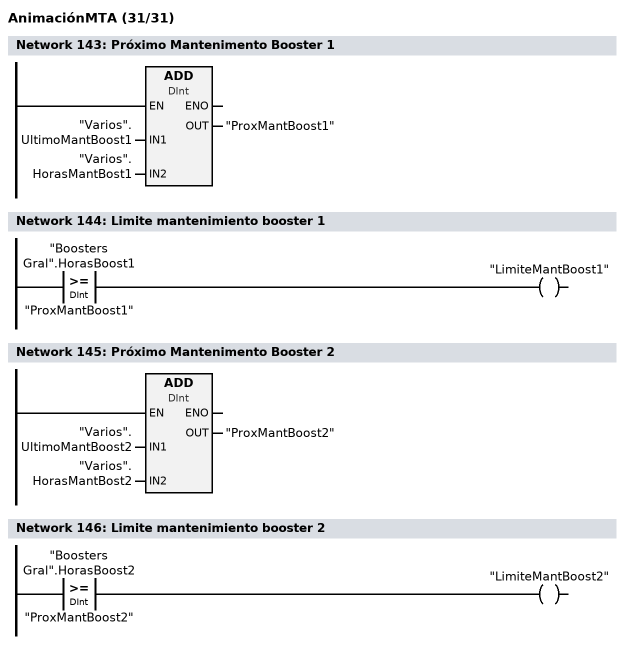
   RUNG wire#powerrail
      { S7_Templates := "SrcType := DInt"; S7_GenerateENO := "TRUE" } Add(in1 := "Varios".UltimoMantBoost1, in2 := "Varios".HorasMantBost1, out => "ProxMantBoost1")
   END_RUNG
   // the same network as SCL:
   "ProxMantBoost1" := "Varios".UltimoMantBoost1 + "Varios".HorasMantBost1;
END_REGION

REGION Network 144: Limite mantenimiento booster 1
   RUNG wire#powerrail
      { S7_Templates := "SrcType := DInt" } GE_Contact(in1 := "Boosters Gral".HorasBoost1, in2 := "ProxMantBoost1")
      Coil( "LimiteMantBoost1" )
   END_RUNG
   // the same network as SCL:
   "LimiteMantBoost1" := "Boosters Gral".HorasBoost1 >= "ProxMantBoost1";
END_REGION

REGION Network 145: Próximo Mantenimento Booster 2
   RUNG wire#powerrail
      { S7_Templates := "SrcType := DInt"; S7_GenerateENO := "TRUE" } Add(in1 := "Varios".UltimoMantBoost2, in2 := "Varios".HorasMantBost2, out => "ProxMantBoost2")
   END_RUNG
   // the same network as SCL:
   "ProxMantBoost2" := "Varios".UltimoMantBoost2 + "Varios".HorasMantBost2;
END_REGION

REGION Network 146: Limite mantenimiento booster 2
   RUNG wire#powerrail
      { S7_Templates := "SrcType := DInt" } GE_Contact(in1 := "Boosters Gral".HorasBoost2, in2 := "ProxMantBoost2")
      Coil( "LimiteMantBoost2" )
   END_RUNG
   // the same network as SCL:
   "LimiteMantBoost2" := "Boosters Gral".HorasBoost2 >= "ProxMantBoost2";
END_REGION
END_FUNCTION

FUNCTION "Motores-PanelMTA" : Void   // FC3, LAD
{ S7_Optimized_Access := 'FALSE' }
VERSION : 0.1
BEGIN

REGION Network 1: Comandos desde Panel para MP010 - Bomba Principal Ch. Soplado
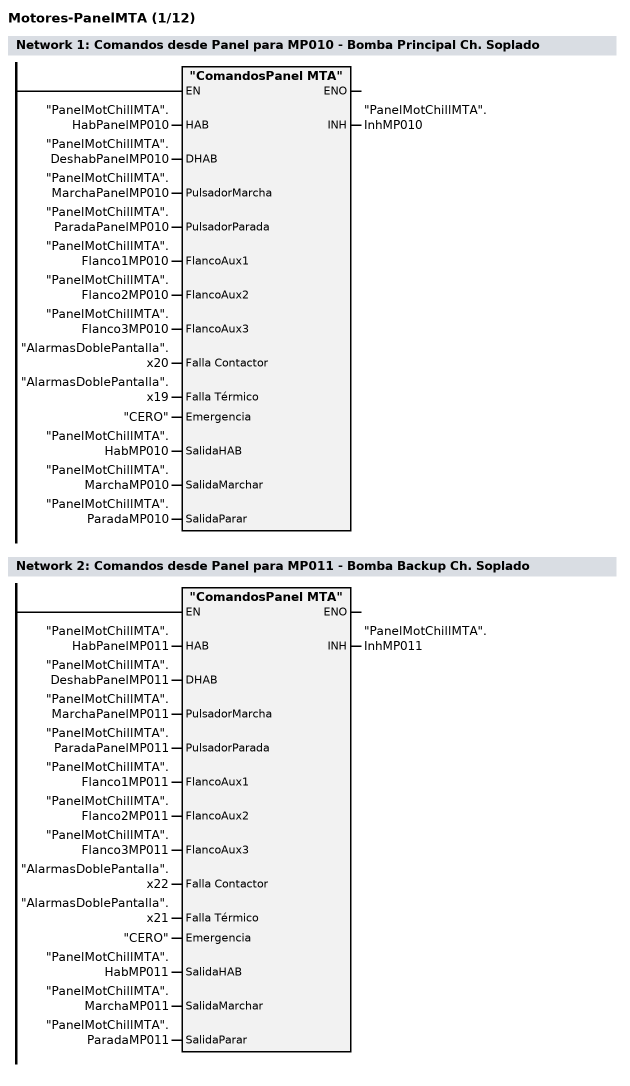
   RUNG wire#powerrail
      "ComandosPanel MTA"(HAB := "PanelMotChillMTA".HabPanelMP010, DHAB := "PanelMotChillMTA".DeshabPanelMP010, PulsadorMarcha := "PanelMotChillMTA".MarchaPanelMP010, PulsadorParada := "PanelMotChillMTA".ParadaPanelMP010, FlancoAux1 := "PanelMotChillMTA".Flanco1MP010, FlancoAux2 := "PanelMotChillMTA".Flanco2MP010, FlancoAux3 := "PanelMotChillMTA".Flanco3MP010, "Falla Contactor" := "AlarmasDoblePantalla".x20, "Falla Térmico" := "AlarmasDoblePantalla".x19, Emergencia := "CERO", INH => "PanelMotChillMTA".InhMP010, SalidaHAB := "PanelMotChillMTA".HabMP010, SalidaMarchar := "PanelMotChillMTA".MarchaMP010, SalidaParar := "PanelMotChillMTA".ParadaMP010)
   END_RUNG
   // the same network as SCL:
   "ComandosPanel MTA"(HAB := "PanelMotChillMTA".HabPanelMP010,
                       DHAB := "PanelMotChillMTA".DeshabPanelMP010,
                       PulsadorMarcha := "PanelMotChillMTA".MarchaPanelMP010,
                       PulsadorParada := "PanelMotChillMTA".ParadaPanelMP010,
                       FlancoAux1 := "PanelMotChillMTA".Flanco1MP010,
                       FlancoAux2 := "PanelMotChillMTA".Flanco2MP010,
                       FlancoAux3 := "PanelMotChillMTA".Flanco3MP010,
                       "Falla Contactor" := "AlarmasDoblePantalla".x20,
                       "Falla Térmico" := "AlarmasDoblePantalla".x19,
                       Emergencia := "CERO",
                       SalidaHAB := "PanelMotChillMTA".HabMP010,
                       SalidaMarchar := "PanelMotChillMTA".MarchaMP010,
                       SalidaParar := "PanelMotChillMTA".ParadaMP010,
                       INH => "PanelMotChillMTA".InhMP010);
END_REGION

REGION Network 2: Comandos desde Panel para MP011 - Bomba Backup Ch. Soplado
   RUNG wire#powerrail
      "ComandosPanel MTA"(HAB := "PanelMotChillMTA".HabPanelMP011, DHAB := "PanelMotChillMTA".DeshabPanelMP011, PulsadorMarcha := "PanelMotChillMTA".MarchaPanelMP011, PulsadorParada := "PanelMotChillMTA".ParadaPanelMP011, FlancoAux1 := "PanelMotChillMTA".Flanco1MP011, FlancoAux2 := "PanelMotChillMTA".Flanco2MP011, FlancoAux3 := "PanelMotChillMTA".Flanco3MP011, "Falla Contactor" := "AlarmasDoblePantalla".x22, "Falla Térmico" := "AlarmasDoblePantalla".x21, Emergencia := "CERO", INH => "PanelMotChillMTA".InhMP011, SalidaHAB := "PanelMotChillMTA".HabMP011, SalidaMarchar := "PanelMotChillMTA".MarchaMP011, SalidaParar := "PanelMotChillMTA".ParadaMP011)
   END_RUNG
   // the same network as SCL:
   "ComandosPanel MTA"(HAB := "PanelMotChillMTA".HabPanelMP011,
                       DHAB := "PanelMotChillMTA".DeshabPanelMP011,
                       PulsadorMarcha := "PanelMotChillMTA".MarchaPanelMP011,
                       PulsadorParada := "PanelMotChillMTA".ParadaPanelMP011,
                       FlancoAux1 := "PanelMotChillMTA".Flanco1MP011,
                       FlancoAux2 := "PanelMotChillMTA".Flanco2MP011,
                       FlancoAux3 := "PanelMotChillMTA".Flanco3MP011,
                       "Falla Contactor" := "AlarmasDoblePantalla".x22,
                       "Falla Térmico" := "AlarmasDoblePantalla".x21,
                       Emergencia := "CERO",
                       SalidaHAB := "PanelMotChillMTA".HabMP011,
                       SalidaMarchar := "PanelMotChillMTA".MarchaMP011,
                       SalidaParar := "PanelMotChillMTA".ParadaMP011,
                       INH => "PanelMotChillMTA".InhMP011);
END_REGION

REGION Network 3: Comandos desde Panel para MP012 - Bomba Principal Ch. Envasado
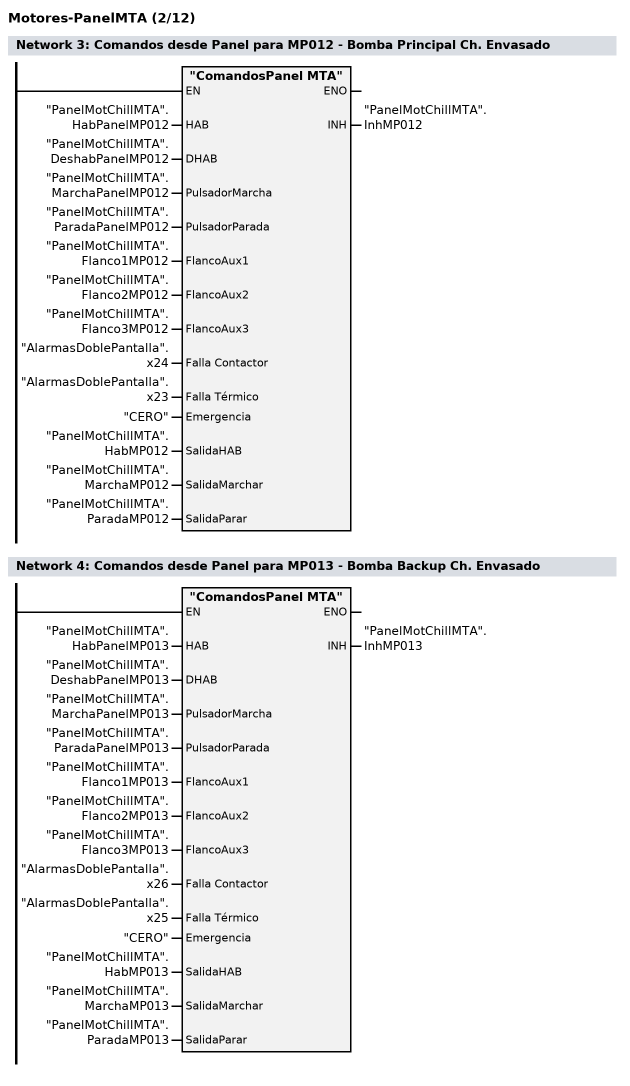
   RUNG wire#powerrail
      "ComandosPanel MTA"(HAB := "PanelMotChillMTA".HabPanelMP012, DHAB := "PanelMotChillMTA".DeshabPanelMP012, PulsadorMarcha := "PanelMotChillMTA".MarchaPanelMP012, PulsadorParada := "PanelMotChillMTA".ParadaPanelMP012, FlancoAux1 := "PanelMotChillMTA".Flanco1MP012, FlancoAux2 := "PanelMotChillMTA".Flanco2MP012, FlancoAux3 := "PanelMotChillMTA".Flanco3MP012, "Falla Contactor" := "AlarmasDoblePantalla".x24, "Falla Térmico" := "AlarmasDoblePantalla".x23, Emergencia := "CERO", INH => "PanelMotChillMTA".InhMP012, SalidaHAB := "PanelMotChillMTA".HabMP012, SalidaMarchar := "PanelMotChillMTA".MarchaMP012, SalidaParar := "PanelMotChillMTA".ParadaMP012)
   END_RUNG
   // the same network as SCL:
   "ComandosPanel MTA"(HAB := "PanelMotChillMTA".HabPanelMP012,
                       DHAB := "PanelMotChillMTA".DeshabPanelMP012,
                       PulsadorMarcha := "PanelMotChillMTA".MarchaPanelMP012,
                       PulsadorParada := "PanelMotChillMTA".ParadaPanelMP012,
                       FlancoAux1 := "PanelMotChillMTA".Flanco1MP012,
                       FlancoAux2 := "PanelMotChillMTA".Flanco2MP012,
                       FlancoAux3 := "PanelMotChillMTA".Flanco3MP012,
                       "Falla Contactor" := "AlarmasDoblePantalla".x24,
                       "Falla Térmico" := "AlarmasDoblePantalla".x23,
                       Emergencia := "CERO",
                       SalidaHAB := "PanelMotChillMTA".HabMP012,
                       SalidaMarchar := "PanelMotChillMTA".MarchaMP012,
                       SalidaParar := "PanelMotChillMTA".ParadaMP012,
                       INH => "PanelMotChillMTA".InhMP012);
END_REGION

REGION Network 4: Comandos desde Panel para MP013 - Bomba Backup Ch. Envasado
   RUNG wire#powerrail
      "ComandosPanel MTA"(HAB := "PanelMotChillMTA".HabPanelMP013, DHAB := "PanelMotChillMTA".DeshabPanelMP013, PulsadorMarcha := "PanelMotChillMTA".MarchaPanelMP013, PulsadorParada := "PanelMotChillMTA".ParadaPanelMP013, FlancoAux1 := "PanelMotChillMTA".Flanco1MP013, FlancoAux2 := "PanelMotChillMTA".Flanco2MP013, FlancoAux3 := "PanelMotChillMTA".Flanco3MP013, "Falla Contactor" := "AlarmasDoblePantalla".x26, "Falla Térmico" := "AlarmasDoblePantalla".x25, Emergencia := "CERO", INH => "PanelMotChillMTA".InhMP013, SalidaHAB := "PanelMotChillMTA".HabMP013, SalidaMarchar := "PanelMotChillMTA".MarchaMP013, SalidaParar := "PanelMotChillMTA".ParadaMP013)
   END_RUNG
   // the same network as SCL:
   "ComandosPanel MTA"(HAB := "PanelMotChillMTA".HabPanelMP013,
                       DHAB := "PanelMotChillMTA".DeshabPanelMP013,
                       PulsadorMarcha := "PanelMotChillMTA".MarchaPanelMP013,
                       PulsadorParada := "PanelMotChillMTA".ParadaPanelMP013,
                       FlancoAux1 := "PanelMotChillMTA".Flanco1MP013,
                       FlancoAux2 := "PanelMotChillMTA".Flanco2MP013,
                       FlancoAux3 := "PanelMotChillMTA".Flanco3MP013,
                       "Falla Contactor" := "AlarmasDoblePantalla".x26,
                       "Falla Térmico" := "AlarmasDoblePantalla".x25,
                       Emergencia := "CERO",
                       SalidaHAB := "PanelMotChillMTA".HabMP013,
                       SalidaMarchar := "PanelMotChillMTA".MarchaMP013,
                       SalidaParar := "PanelMotChillMTA".ParadaMP013,
                       INH => "PanelMotChillMTA".InhMP013);
END_REGION

REGION Network 5: Comandos desde Panel para MP018 - Bomba 1 Torres de enfriamiento Chillers
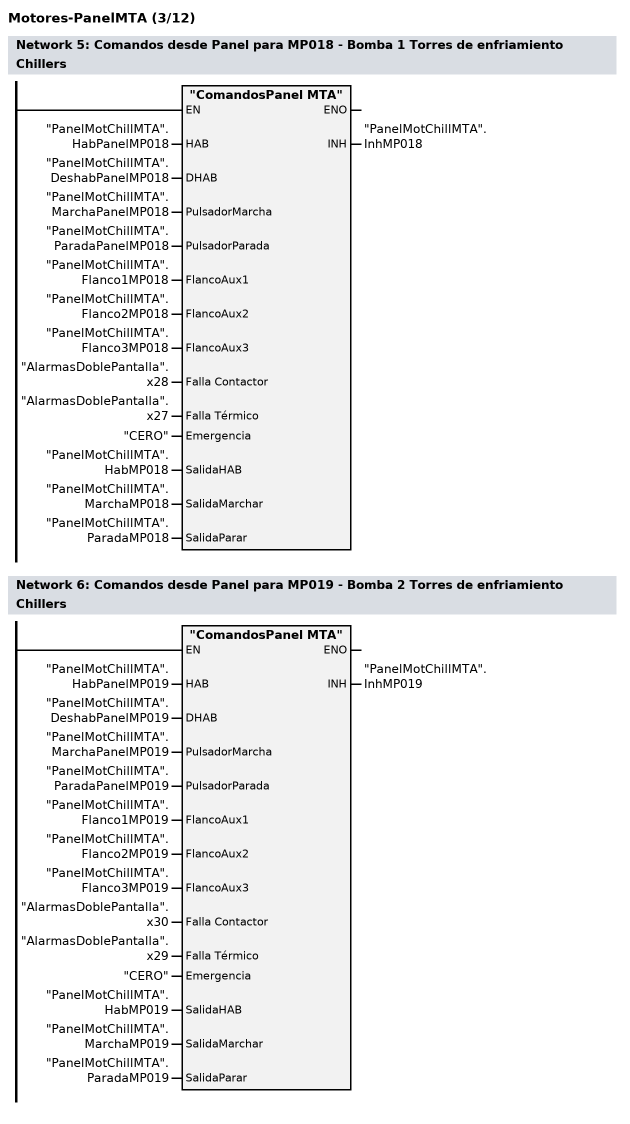
   RUNG wire#powerrail
      "ComandosPanel MTA"(HAB := "PanelMotChillMTA".HabPanelMP018, DHAB := "PanelMotChillMTA".DeshabPanelMP018, PulsadorMarcha := "PanelMotChillMTA".MarchaPanelMP018, PulsadorParada := "PanelMotChillMTA".ParadaPanelMP018, FlancoAux1 := "PanelMotChillMTA".Flanco1MP018, FlancoAux2 := "PanelMotChillMTA".Flanco2MP018, FlancoAux3 := "PanelMotChillMTA".Flanco3MP018, "Falla Contactor" := "AlarmasDoblePantalla".x28, "Falla Térmico" := "AlarmasDoblePantalla".x27, Emergencia := "CERO", SalidaHAB := "PanelMotChillMTA".HabMP018, SalidaMarchar := "PanelMotChillMTA".MarchaMP018, SalidaParar := "PanelMotChillMTA".ParadaMP018, INH => "PanelMotChillMTA".InhMP018)
   END_RUNG
   // the same network as SCL:
   "ComandosPanel MTA"(HAB := "PanelMotChillMTA".HabPanelMP018,
                       DHAB := "PanelMotChillMTA".DeshabPanelMP018,
                       PulsadorMarcha := "PanelMotChillMTA".MarchaPanelMP018,
                       PulsadorParada := "PanelMotChillMTA".ParadaPanelMP018,
                       FlancoAux1 := "PanelMotChillMTA".Flanco1MP018,
                       FlancoAux2 := "PanelMotChillMTA".Flanco2MP018,
                       FlancoAux3 := "PanelMotChillMTA".Flanco3MP018,
                       "Falla Contactor" := "AlarmasDoblePantalla".x28,
                       "Falla Térmico" := "AlarmasDoblePantalla".x27,
                       Emergencia := "CERO",
                       SalidaHAB := "PanelMotChillMTA".HabMP018,
                       SalidaMarchar := "PanelMotChillMTA".MarchaMP018,
                       SalidaParar := "PanelMotChillMTA".ParadaMP018,
                       INH => "PanelMotChillMTA".InhMP018);
END_REGION

REGION Network 6: Comandos desde Panel para MP019 - Bomba 2 Torres de enfriamiento Chillers
   RUNG wire#powerrail
      "ComandosPanel MTA"(HAB := "PanelMotChillMTA".HabPanelMP019, DHAB := "PanelMotChillMTA".DeshabPanelMP019, PulsadorMarcha := "PanelMotChillMTA".MarchaPanelMP019, PulsadorParada := "PanelMotChillMTA".ParadaPanelMP019, FlancoAux1 := "PanelMotChillMTA".Flanco1MP019, FlancoAux2 := "PanelMotChillMTA".Flanco2MP019, FlancoAux3 := "PanelMotChillMTA".Flanco3MP019, "Falla Contactor" := "AlarmasDoblePantalla".x30, "Falla Térmico" := "AlarmasDoblePantalla".x29, Emergencia := "CERO", SalidaHAB := "PanelMotChillMTA".HabMP019, SalidaMarchar := "PanelMotChillMTA".MarchaMP019, SalidaParar := "PanelMotChillMTA".ParadaMP019, INH => "PanelMotChillMTA".InhMP019)
   END_RUNG
   // the same network as SCL:
   "ComandosPanel MTA"(HAB := "PanelMotChillMTA".HabPanelMP019,
                       DHAB := "PanelMotChillMTA".DeshabPanelMP019,
                       PulsadorMarcha := "PanelMotChillMTA".MarchaPanelMP019,
                       PulsadorParada := "PanelMotChillMTA".ParadaPanelMP019,
                       FlancoAux1 := "PanelMotChillMTA".Flanco1MP019,
                       FlancoAux2 := "PanelMotChillMTA".Flanco2MP019,
                       FlancoAux3 := "PanelMotChillMTA".Flanco3MP019,
                       "Falla Contactor" := "AlarmasDoblePantalla".x30,
                       "Falla Térmico" := "AlarmasDoblePantalla".x29,
                       Emergencia := "CERO",
                       SalidaHAB := "PanelMotChillMTA".HabMP019,
                       SalidaMarchar := "PanelMotChillMTA".MarchaMP019,
                       SalidaParar := "PanelMotChillMTA".ParadaMP019,
                       INH => "PanelMotChillMTA".InhMP019);
END_REGION

REGION Network 7: Comandos desde Panel para MT007 - Bomba Soplado L1
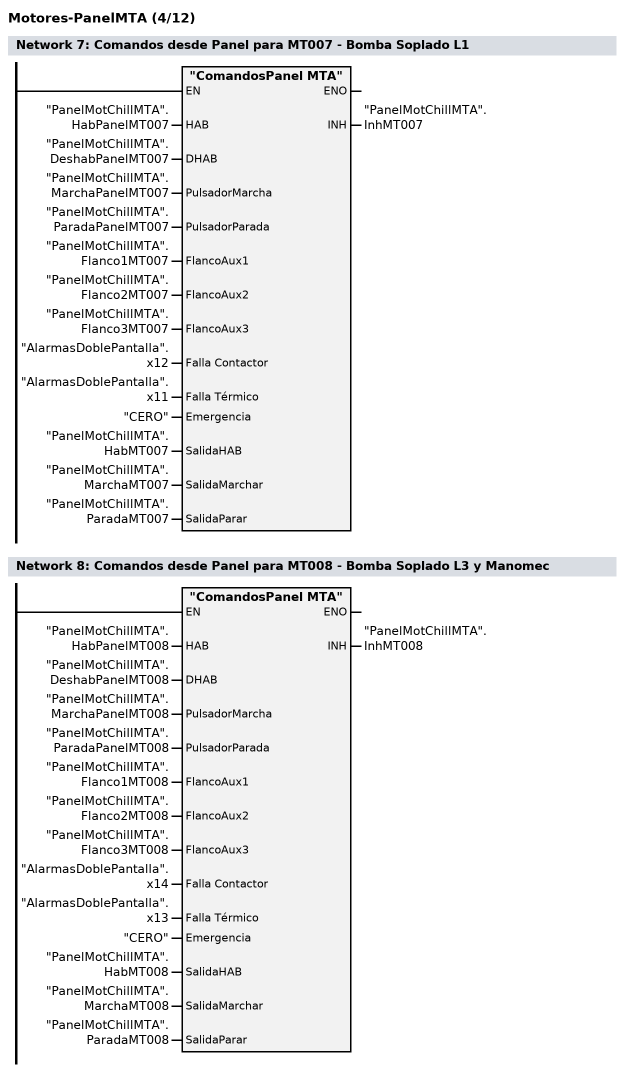
   RUNG wire#powerrail
      "ComandosPanel MTA"(HAB := "PanelMotChillMTA".HabPanelMT007, DHAB := "PanelMotChillMTA".DeshabPanelMT007, PulsadorMarcha := "PanelMotChillMTA".MarchaPanelMT007, PulsadorParada := "PanelMotChillMTA".ParadaPanelMT007, FlancoAux1 := "PanelMotChillMTA".Flanco1MT007, FlancoAux2 := "PanelMotChillMTA".Flanco2MT007, FlancoAux3 := "PanelMotChillMTA".Flanco3MT007, "Falla Contactor" := "AlarmasDoblePantalla".x12, "Falla Térmico" := "AlarmasDoblePantalla".x11, Emergencia := "CERO", INH => "PanelMotChillMTA".InhMT007, SalidaHAB := "PanelMotChillMTA".HabMT007, SalidaMarchar := "PanelMotChillMTA".MarchaMT007, SalidaParar := "PanelMotChillMTA".ParadaMT007)
   END_RUNG
   // the same network as SCL:
   "ComandosPanel MTA"(HAB := "PanelMotChillMTA".HabPanelMT007,
                       DHAB := "PanelMotChillMTA".DeshabPanelMT007,
                       PulsadorMarcha := "PanelMotChillMTA".MarchaPanelMT007,
                       PulsadorParada := "PanelMotChillMTA".ParadaPanelMT007,
                       FlancoAux1 := "PanelMotChillMTA".Flanco1MT007,
                       FlancoAux2 := "PanelMotChillMTA".Flanco2MT007,
                       FlancoAux3 := "PanelMotChillMTA".Flanco3MT007,
                       "Falla Contactor" := "AlarmasDoblePantalla".x12,
                       "Falla Térmico" := "AlarmasDoblePantalla".x11,
                       Emergencia := "CERO",
                       SalidaHAB := "PanelMotChillMTA".HabMT007,
                       SalidaMarchar := "PanelMotChillMTA".MarchaMT007,
                       SalidaParar := "PanelMotChillMTA".ParadaMT007,
                       INH => "PanelMotChillMTA".InhMT007);
END_REGION

REGION Network 8: Comandos desde Panel para MT008 - Bomba Soplado L3 y Manomec
   RUNG wire#powerrail
      "ComandosPanel MTA"(HAB := "PanelMotChillMTA".HabPanelMT008, DHAB := "PanelMotChillMTA".DeshabPanelMT008, PulsadorMarcha := "PanelMotChillMTA".MarchaPanelMT008, PulsadorParada := "PanelMotChillMTA".ParadaPanelMT008, FlancoAux1 := "PanelMotChillMTA".Flanco1MT008, FlancoAux2 := "PanelMotChillMTA".Flanco2MT008, FlancoAux3 := "PanelMotChillMTA".Flanco3MT008, "Falla Contactor" := "AlarmasDoblePantalla".x14, "Falla Térmico" := "AlarmasDoblePantalla".x13, Emergencia := "CERO", INH => "PanelMotChillMTA".InhMT008, SalidaHAB := "PanelMotChillMTA".HabMT008, SalidaMarchar := "PanelMotChillMTA".MarchaMT008, SalidaParar := "PanelMotChillMTA".ParadaMT008)
   END_RUNG
   // the same network as SCL:
   "ComandosPanel MTA"(HAB := "PanelMotChillMTA".HabPanelMT008,
                       DHAB := "PanelMotChillMTA".DeshabPanelMT008,
                       PulsadorMarcha := "PanelMotChillMTA".MarchaPanelMT008,
                       PulsadorParada := "PanelMotChillMTA".ParadaPanelMT008,
                       FlancoAux1 := "PanelMotChillMTA".Flanco1MT008,
                       FlancoAux2 := "PanelMotChillMTA".Flanco2MT008,
                       FlancoAux3 := "PanelMotChillMTA".Flanco3MT008,
                       "Falla Contactor" := "AlarmasDoblePantalla".x14,
                       "Falla Térmico" := "AlarmasDoblePantalla".x13,
                       Emergencia := "CERO",
                       SalidaHAB := "PanelMotChillMTA".HabMT008,
                       SalidaMarchar := "PanelMotChillMTA".MarchaMT008,
                       SalidaParar := "PanelMotChillMTA".ParadaMT008,
                       INH => "PanelMotChillMTA".InhMT008);
END_REGION

REGION Network 9: Comandos desde Panel para MT009 - Bomba Int. L3 y L5
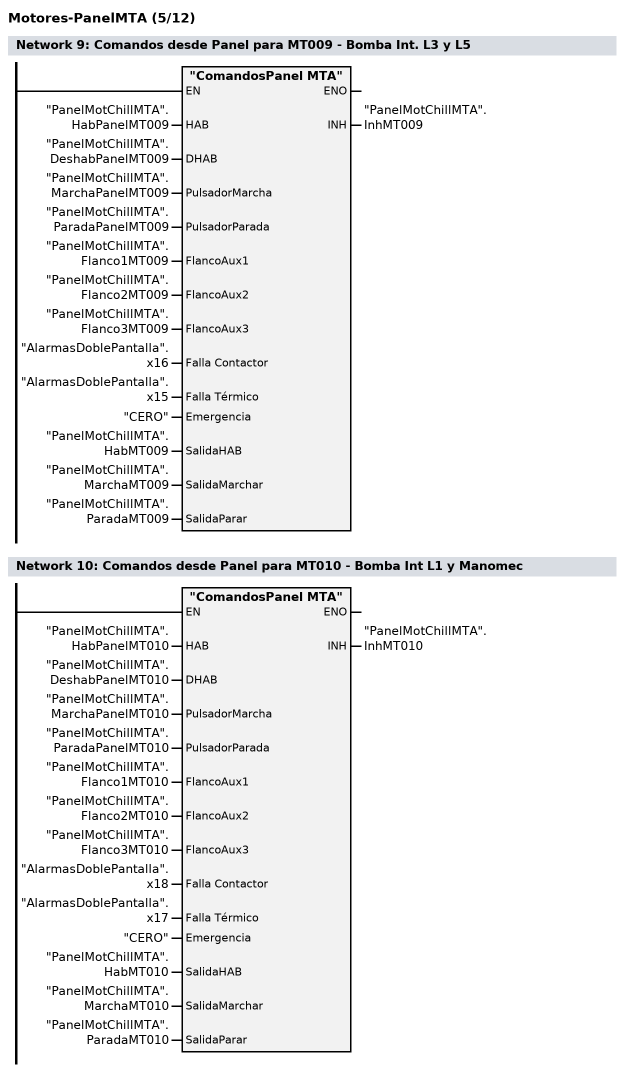
   RUNG wire#powerrail
      "ComandosPanel MTA"(HAB := "PanelMotChillMTA".HabPanelMT009, DHAB := "PanelMotChillMTA".DeshabPanelMT009, PulsadorMarcha := "PanelMotChillMTA".MarchaPanelMT009, PulsadorParada := "PanelMotChillMTA".ParadaPanelMT009, FlancoAux1 := "PanelMotChillMTA".Flanco1MT009, FlancoAux2 := "PanelMotChillMTA".Flanco2MT009, FlancoAux3 := "PanelMotChillMTA".Flanco3MT009, "Falla Contactor" := "AlarmasDoblePantalla".x16, "Falla Térmico" := "AlarmasDoblePantalla".x15, Emergencia := "CERO", INH => "PanelMotChillMTA".InhMT009, SalidaHAB := "PanelMotChillMTA".HabMT009, SalidaMarchar := "PanelMotChillMTA".MarchaMT009, SalidaParar := "PanelMotChillMTA".ParadaMT009)
   END_RUNG
   // the same network as SCL:
   "ComandosPanel MTA"(HAB := "PanelMotChillMTA".HabPanelMT009,
                       DHAB := "PanelMotChillMTA".DeshabPanelMT009,
                       PulsadorMarcha := "PanelMotChillMTA".MarchaPanelMT009,
                       PulsadorParada := "PanelMotChillMTA".ParadaPanelMT009,
                       FlancoAux1 := "PanelMotChillMTA".Flanco1MT009,
                       FlancoAux2 := "PanelMotChillMTA".Flanco2MT009,
                       FlancoAux3 := "PanelMotChillMTA".Flanco3MT009,
                       "Falla Contactor" := "AlarmasDoblePantalla".x16,
                       "Falla Térmico" := "AlarmasDoblePantalla".x15,
                       Emergencia := "CERO",
                       SalidaHAB := "PanelMotChillMTA".HabMT009,
                       SalidaMarchar := "PanelMotChillMTA".MarchaMT009,
                       SalidaParar := "PanelMotChillMTA".ParadaMT009,
                       INH => "PanelMotChillMTA".InhMT009);
END_REGION

REGION Network 10: Comandos desde Panel para MT010 - Bomba Int L1 y Manomec
   RUNG wire#powerrail
      "ComandosPanel MTA"(HAB := "PanelMotChillMTA".HabPanelMT010, DHAB := "PanelMotChillMTA".DeshabPanelMT010, PulsadorMarcha := "PanelMotChillMTA".MarchaPanelMT010, PulsadorParada := "PanelMotChillMTA".ParadaPanelMT010, FlancoAux1 := "PanelMotChillMTA".Flanco1MT010, FlancoAux2 := "PanelMotChillMTA".Flanco2MT010, FlancoAux3 := "PanelMotChillMTA".Flanco3MT010, "Falla Contactor" := "AlarmasDoblePantalla".x18, "Falla Térmico" := "AlarmasDoblePantalla".x17, Emergencia := "CERO", INH => "PanelMotChillMTA".InhMT010, SalidaHAB := "PanelMotChillMTA".HabMT010, SalidaMarchar := "PanelMotChillMTA".MarchaMT010, SalidaParar := "PanelMotChillMTA".ParadaMT010)
   END_RUNG
   // the same network as SCL:
   "ComandosPanel MTA"(HAB := "PanelMotChillMTA".HabPanelMT010,
                       DHAB := "PanelMotChillMTA".DeshabPanelMT010,
                       PulsadorMarcha := "PanelMotChillMTA".MarchaPanelMT010,
                       PulsadorParada := "PanelMotChillMTA".ParadaPanelMT010,
                       FlancoAux1 := "PanelMotChillMTA".Flanco1MT010,
                       FlancoAux2 := "PanelMotChillMTA".Flanco2MT010,
                       FlancoAux3 := "PanelMotChillMTA".Flanco3MT010,
                       "Falla Contactor" := "AlarmasDoblePantalla".x18,
                       "Falla Térmico" := "AlarmasDoblePantalla".x17,
                       Emergencia := "CERO",
                       SalidaHAB := "PanelMotChillMTA".HabMT010,
                       SalidaMarchar := "PanelMotChillMTA".MarchaMT010,
                       SalidaParar := "PanelMotChillMTA".ParadaMT010,
                       INH => "PanelMotChillMTA".InhMT010);
END_REGION

REGION Network 11: Comandos desde Panel para V001 - Ventilador 1 Torres de enfriamiento Chillers
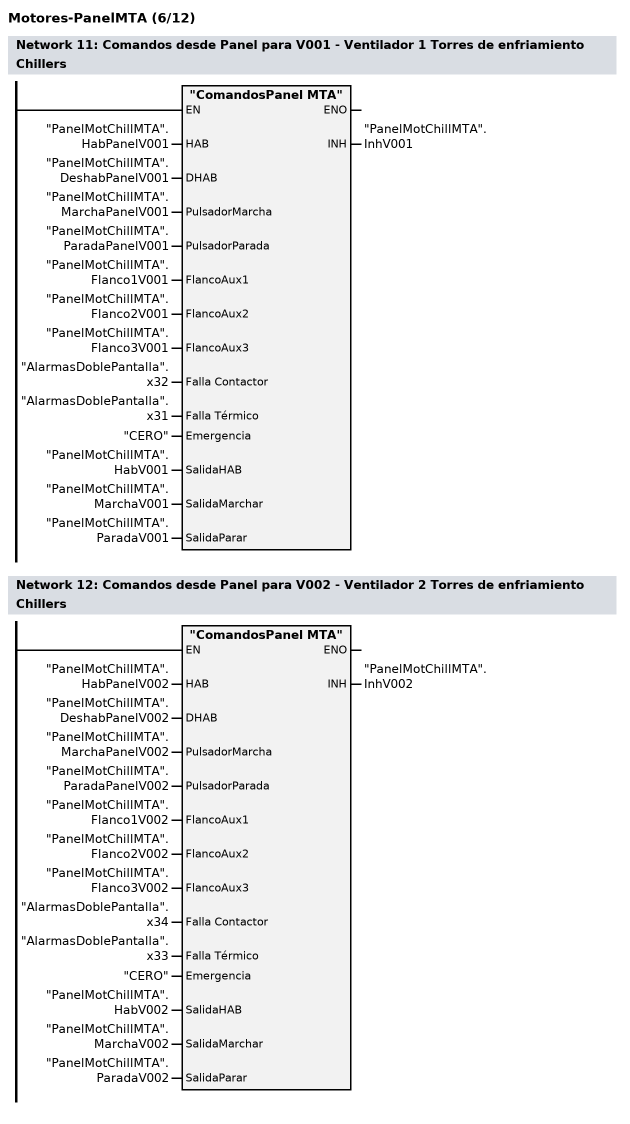
   RUNG wire#powerrail
      "ComandosPanel MTA"(HAB := "PanelMotChillMTA".HabPanelV001, DHAB := "PanelMotChillMTA".DeshabPanelV001, PulsadorMarcha := "PanelMotChillMTA".MarchaPanelV001, PulsadorParada := "PanelMotChillMTA".ParadaPanelV001, FlancoAux1 := "PanelMotChillMTA".Flanco1V001, FlancoAux2 := "PanelMotChillMTA".Flanco2V001, FlancoAux3 := "PanelMotChillMTA".Flanco3V001, "Falla Contactor" := "AlarmasDoblePantalla".x32, "Falla Térmico" := "AlarmasDoblePantalla".x31, Emergencia := "CERO", SalidaHAB := "PanelMotChillMTA".HabV001, SalidaMarchar := "PanelMotChillMTA".MarchaV001, SalidaParar := "PanelMotChillMTA".ParadaV001, INH => "PanelMotChillMTA".InhV001)
   END_RUNG
   // the same network as SCL:
   "ComandosPanel MTA"(HAB := "PanelMotChillMTA".HabPanelV001,
                       DHAB := "PanelMotChillMTA".DeshabPanelV001,
                       PulsadorMarcha := "PanelMotChillMTA".MarchaPanelV001,
                       PulsadorParada := "PanelMotChillMTA".ParadaPanelV001,
                       FlancoAux1 := "PanelMotChillMTA".Flanco1V001,
                       FlancoAux2 := "PanelMotChillMTA".Flanco2V001,
                       FlancoAux3 := "PanelMotChillMTA".Flanco3V001,
                       "Falla Contactor" := "AlarmasDoblePantalla".x32,
                       "Falla Térmico" := "AlarmasDoblePantalla".x31,
                       Emergencia := "CERO",
                       SalidaHAB := "PanelMotChillMTA".HabV001,
                       SalidaMarchar := "PanelMotChillMTA".MarchaV001,
                       SalidaParar := "PanelMotChillMTA".ParadaV001,
                       INH => "PanelMotChillMTA".InhV001);
END_REGION

REGION Network 12: Comandos desde Panel para V002 - Ventilador 2 Torres de enfriamiento Chillers
   RUNG wire#powerrail
      "ComandosPanel MTA"(HAB := "PanelMotChillMTA".HabPanelV002, DHAB := "PanelMotChillMTA".DeshabPanelV002, PulsadorMarcha := "PanelMotChillMTA".MarchaPanelV002, PulsadorParada := "PanelMotChillMTA".ParadaPanelV002, FlancoAux1 := "PanelMotChillMTA".Flanco1V002, FlancoAux2 := "PanelMotChillMTA".Flanco2V002, FlancoAux3 := "PanelMotChillMTA".Flanco3V002, "Falla Contactor" := "AlarmasDoblePantalla".x34, "Falla Térmico" := "AlarmasDoblePantalla".x33, Emergencia := "CERO", SalidaHAB := "PanelMotChillMTA".HabV002, SalidaMarchar := "PanelMotChillMTA".MarchaV002, SalidaParar := "PanelMotChillMTA".ParadaV002, INH => "PanelMotChillMTA".InhV002)
   END_RUNG
   // the same network as SCL:
   "ComandosPanel MTA"(HAB := "PanelMotChillMTA".HabPanelV002,
                       DHAB := "PanelMotChillMTA".DeshabPanelV002,
                       PulsadorMarcha := "PanelMotChillMTA".MarchaPanelV002,
                       PulsadorParada := "PanelMotChillMTA".ParadaPanelV002,
                       FlancoAux1 := "PanelMotChillMTA".Flanco1V002,
                       FlancoAux2 := "PanelMotChillMTA".Flanco2V002,
                       FlancoAux3 := "PanelMotChillMTA".Flanco3V002,
                       "Falla Contactor" := "AlarmasDoblePantalla".x34,
                       "Falla Térmico" := "AlarmasDoblePantalla".x33,
                       Emergencia := "CERO",
                       SalidaHAB := "PanelMotChillMTA".HabV002,
                       SalidaMarchar := "PanelMotChillMTA".MarchaV002,
                       SalidaParar := "PanelMotChillMTA".ParadaV002,
                       INH => "PanelMotChillMTA".InhV002);
END_REGION

REGION Network 13: Comandos desde Panel para V003 - Ventilador 3 Torres de enfriamiento Chillers
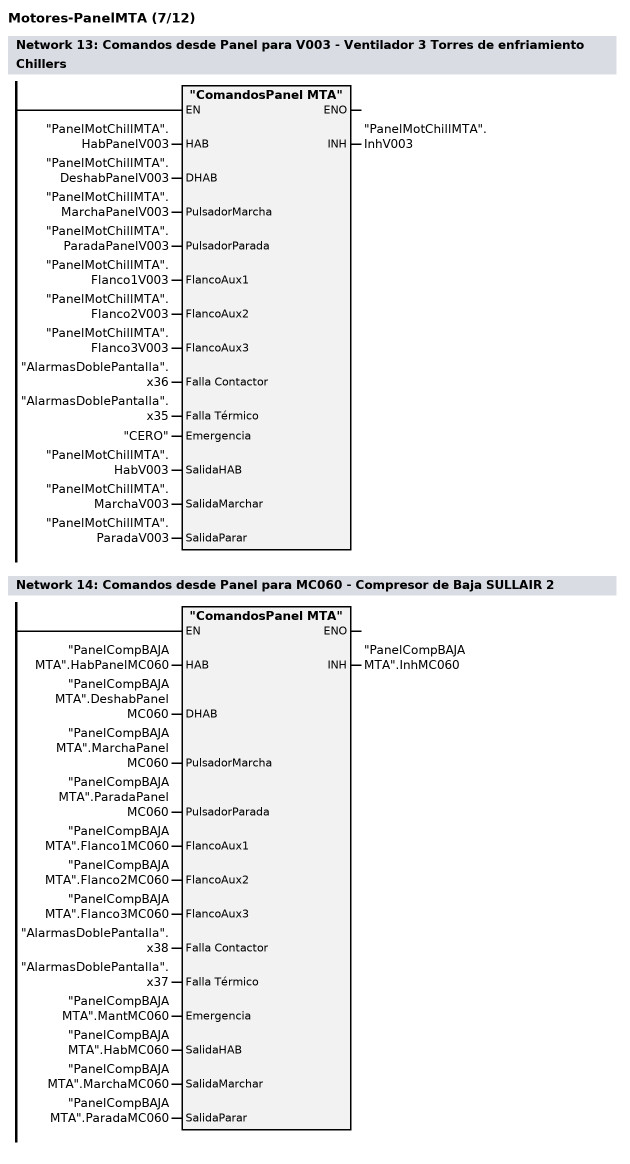
   RUNG wire#powerrail
      "ComandosPanel MTA"(HAB := "PanelMotChillMTA".HabPanelV003, DHAB := "PanelMotChillMTA".DeshabPanelV003, PulsadorMarcha := "PanelMotChillMTA".MarchaPanelV003, PulsadorParada := "PanelMotChillMTA".ParadaPanelV003, FlancoAux1 := "PanelMotChillMTA".Flanco1V003, FlancoAux2 := "PanelMotChillMTA".Flanco2V003, FlancoAux3 := "PanelMotChillMTA".Flanco3V003, "Falla Contactor" := "AlarmasDoblePantalla".x36, "Falla Térmico" := "AlarmasDoblePantalla".x35, Emergencia := "CERO", SalidaHAB := "PanelMotChillMTA".HabV003, SalidaMarchar := "PanelMotChillMTA".MarchaV003, SalidaParar := "PanelMotChillMTA".ParadaV003, INH => "PanelMotChillMTA".InhV003)
   END_RUNG
   // the same network as SCL:
   "ComandosPanel MTA"(HAB := "PanelMotChillMTA".HabPanelV003,
                       DHAB := "PanelMotChillMTA".DeshabPanelV003,
                       PulsadorMarcha := "PanelMotChillMTA".MarchaPanelV003,
                       PulsadorParada := "PanelMotChillMTA".ParadaPanelV003,
                       FlancoAux1 := "PanelMotChillMTA".Flanco1V003,
                       FlancoAux2 := "PanelMotChillMTA".Flanco2V003,
                       FlancoAux3 := "PanelMotChillMTA".Flanco3V003,
                       "Falla Contactor" := "AlarmasDoblePantalla".x36,
                       "Falla Térmico" := "AlarmasDoblePantalla".x35,
                       Emergencia := "CERO",
                       SalidaHAB := "PanelMotChillMTA".HabV003,
                       SalidaMarchar := "PanelMotChillMTA".MarchaV003,
                       SalidaParar := "PanelMotChillMTA".ParadaV003,
                       INH => "PanelMotChillMTA".InhV003);
END_REGION

REGION Network 14: Comandos desde Panel para MC060 - Compresor de Baja SULLAIR 2
   RUNG wire#powerrail
      "ComandosPanel MTA"(HAB := "PanelCompBAJA MTA".HabPanelMC060, DHAB := "PanelCompBAJA MTA".DeshabPanelMC060, PulsadorMarcha := "PanelCompBAJA MTA".MarchaPanelMC060, PulsadorParada := "PanelCompBAJA MTA".ParadaPanelMC060, FlancoAux1 := "PanelCompBAJA MTA".Flanco1MC060, FlancoAux2 := "PanelCompBAJA MTA".Flanco2MC060, FlancoAux3 := "PanelCompBAJA MTA".Flanco3MC060, "Falla Contactor" := "AlarmasDoblePantalla".x38, "Falla Térmico" := "AlarmasDoblePantalla".x37, Emergencia := "PanelCompBAJA MTA".MantMC060, INH => "PanelCompBAJA MTA".InhMC060, SalidaHAB := "PanelCompBAJA MTA".HabMC060, SalidaMarchar := "PanelCompBAJA MTA".MarchaMC060, SalidaParar := "PanelCompBAJA MTA".ParadaMC060)
   END_RUNG
   // the same network as SCL:
   "ComandosPanel MTA"(HAB := "PanelCompBAJA MTA".HabPanelMC060,
                       DHAB := "PanelCompBAJA MTA".DeshabPanelMC060,
                       PulsadorMarcha := "PanelCompBAJA MTA".MarchaPanelMC060,
                       PulsadorParada := "PanelCompBAJA MTA".ParadaPanelMC060,
                       FlancoAux1 := "PanelCompBAJA MTA".Flanco1MC060,
                       FlancoAux2 := "PanelCompBAJA MTA".Flanco2MC060,
                       FlancoAux3 := "PanelCompBAJA MTA".Flanco3MC060,
                       "Falla Contactor" := "AlarmasDoblePantalla".x38,
                       "Falla Térmico" := "AlarmasDoblePantalla".x37,
                       Emergencia := "PanelCompBAJA MTA".MantMC060,
                       SalidaHAB := "PanelCompBAJA MTA".HabMC060,
                       SalidaMarchar := "PanelCompBAJA MTA".MarchaMC060,
                       SalidaParar := "PanelCompBAJA MTA".ParadaMC060,
                       INH => "PanelCompBAJA MTA".InhMC060);
END_REGION

REGION Network 15: Comandos desde Panel para MC061 - Compresor de Baja SULLAIR 1
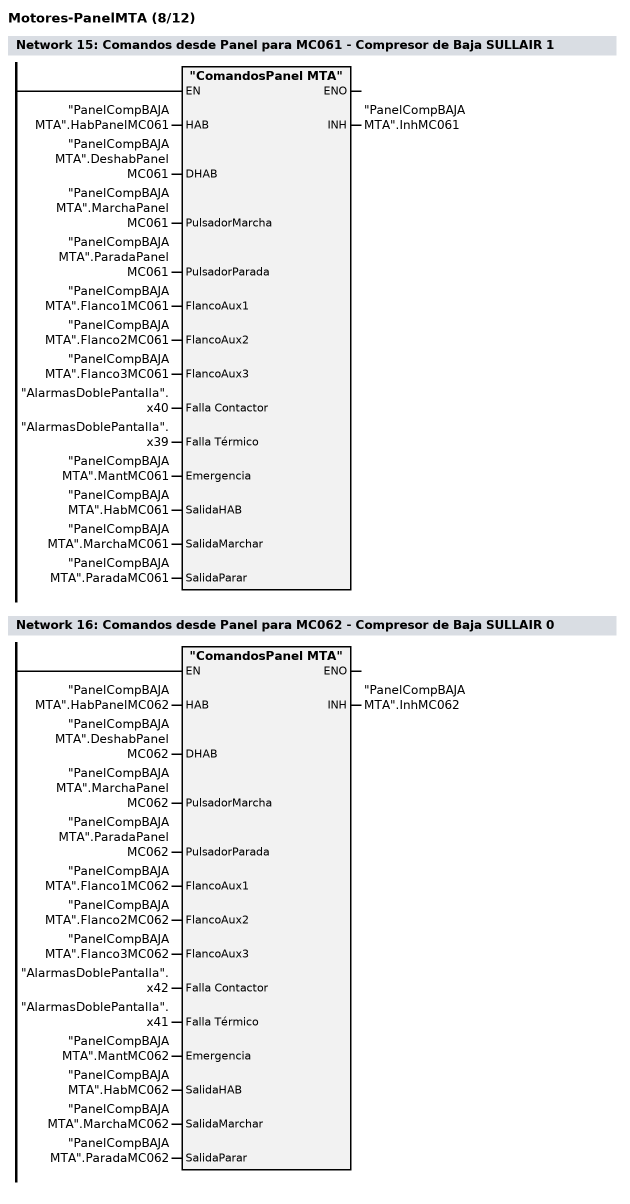
   RUNG wire#powerrail
      "ComandosPanel MTA"(HAB := "PanelCompBAJA MTA".HabPanelMC061, DHAB := "PanelCompBAJA MTA".DeshabPanelMC061, PulsadorMarcha := "PanelCompBAJA MTA".MarchaPanelMC061, PulsadorParada := "PanelCompBAJA MTA".ParadaPanelMC061, FlancoAux1 := "PanelCompBAJA MTA".Flanco1MC061, FlancoAux2 := "PanelCompBAJA MTA".Flanco2MC061, FlancoAux3 := "PanelCompBAJA MTA".Flanco3MC061, "Falla Contactor" := "AlarmasDoblePantalla".x40, "Falla Térmico" := "AlarmasDoblePantalla".x39, Emergencia := "PanelCompBAJA MTA".MantMC061, INH => "PanelCompBAJA MTA".InhMC061, SalidaHAB := "PanelCompBAJA MTA".HabMC061, SalidaMarchar := "PanelCompBAJA MTA".MarchaMC061, SalidaParar := "PanelCompBAJA MTA".ParadaMC061)
   END_RUNG
   // the same network as SCL:
   "ComandosPanel MTA"(HAB := "PanelCompBAJA MTA".HabPanelMC061,
                       DHAB := "PanelCompBAJA MTA".DeshabPanelMC061,
                       PulsadorMarcha := "PanelCompBAJA MTA".MarchaPanelMC061,
                       PulsadorParada := "PanelCompBAJA MTA".ParadaPanelMC061,
                       FlancoAux1 := "PanelCompBAJA MTA".Flanco1MC061,
                       FlancoAux2 := "PanelCompBAJA MTA".Flanco2MC061,
                       FlancoAux3 := "PanelCompBAJA MTA".Flanco3MC061,
                       "Falla Contactor" := "AlarmasDoblePantalla".x40,
                       "Falla Térmico" := "AlarmasDoblePantalla".x39,
                       Emergencia := "PanelCompBAJA MTA".MantMC061,
                       SalidaHAB := "PanelCompBAJA MTA".HabMC061,
                       SalidaMarchar := "PanelCompBAJA MTA".MarchaMC061,
                       SalidaParar := "PanelCompBAJA MTA".ParadaMC061,
                       INH => "PanelCompBAJA MTA".InhMC061);
END_REGION

REGION Network 16: Comandos desde Panel para MC062 - Compresor de Baja SULLAIR 0
   RUNG wire#powerrail
      "ComandosPanel MTA"(HAB := "PanelCompBAJA MTA".HabPanelMC062, DHAB := "PanelCompBAJA MTA".DeshabPanelMC062, PulsadorMarcha := "PanelCompBAJA MTA".MarchaPanelMC062, PulsadorParada := "PanelCompBAJA MTA".ParadaPanelMC062, FlancoAux1 := "PanelCompBAJA MTA".Flanco1MC062, FlancoAux2 := "PanelCompBAJA MTA".Flanco2MC062, FlancoAux3 := "PanelCompBAJA MTA".Flanco3MC062, "Falla Contactor" := "AlarmasDoblePantalla".x42, "Falla Térmico" := "AlarmasDoblePantalla".x41, Emergencia := "PanelCompBAJA MTA".MantMC062, INH => "PanelCompBAJA MTA".InhMC062, SalidaHAB := "PanelCompBAJA MTA".HabMC062, SalidaMarchar := "PanelCompBAJA MTA".MarchaMC062, SalidaParar := "PanelCompBAJA MTA".ParadaMC062)
   END_RUNG
   // the same network as SCL:
   "ComandosPanel MTA"(HAB := "PanelCompBAJA MTA".HabPanelMC062,
                       DHAB := "PanelCompBAJA MTA".DeshabPanelMC062,
                       PulsadorMarcha := "PanelCompBAJA MTA".MarchaPanelMC062,
                       PulsadorParada := "PanelCompBAJA MTA".ParadaPanelMC062,
                       FlancoAux1 := "PanelCompBAJA MTA".Flanco1MC062,
                       FlancoAux2 := "PanelCompBAJA MTA".Flanco2MC062,
                       FlancoAux3 := "PanelCompBAJA MTA".Flanco3MC062,
                       "Falla Contactor" := "AlarmasDoblePantalla".x42,
                       "Falla Térmico" := "AlarmasDoblePantalla".x41,
                       Emergencia := "PanelCompBAJA MTA".MantMC062,
                       SalidaHAB := "PanelCompBAJA MTA".HabMC062,
                       SalidaMarchar := "PanelCompBAJA MTA".MarchaMC062,
                       SalidaParar := "PanelCompBAJA MTA".ParadaMC062,
                       INH => "PanelCompBAJA MTA".InhMC062);
END_REGION

REGION Network 17: Comandos desde Panel para MC063 - Compresor de Baja ATLAS 3
